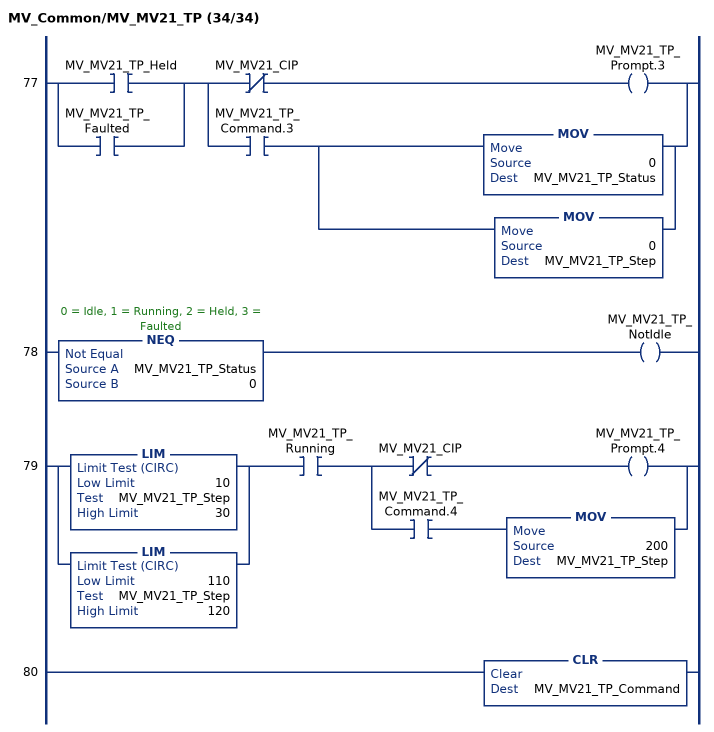
   77: [XIC(MV_MV21_TP_Held) ,XIC(MV_MV21_TP_Faulted) ][XIO(MV_MV21_CIP) OTE(MV_MV21_TP_Prompt.3) ,XIC(MV_MV21_TP_Command.3) [MOV(0,MV_MV21_TP_Status) ,MOV(0,MV_MV21_TP_Step) ] ];
   78: NEQ(MV_MV21_TP_Status,0)OTE(MV_MV21_TP_NotIdle);
   79: [LIM(10,MV_MV21_TP_Step,30) ,LIM(110,MV_MV21_TP_Step,120) ]XIC(MV_MV21_TP_Running)[XIO(MV_MV21_CIP) OTE(MV_MV21_TP_Prompt.4) ,XIC(MV_MV21_TP_Command.4) MOV(200,MV_MV21_TP_Step) ];
   80: CLR(MV_MV21_TP_Command);
END_ROUTINE

ROUTINE MV_MV22_TP   (* ladder *)
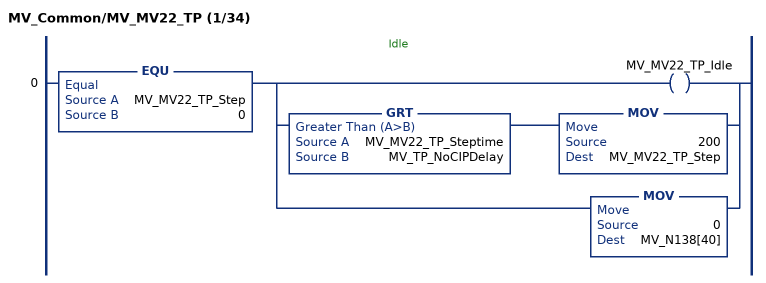
   // Idle
   0: EQU(MV_MV22_TP_Step,0)[OTE(MV_MV22_TP_Idle) ,GRT(MV_MV22_TP_Steptime,MV_TP_NoCIPDelay) MOV(200,MV_MV22_TP_Step) ,MOV(0,MV_N138[40]) ];
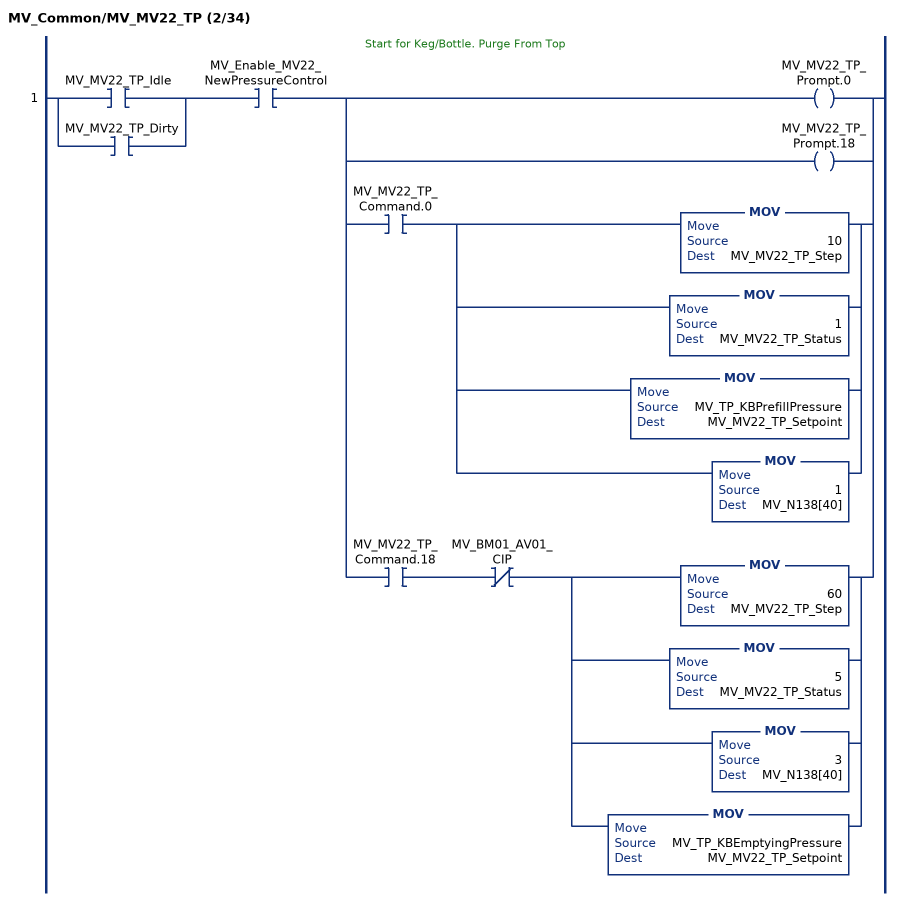
   // Start for Keg/Bottle. Purge From Top
   1: [XIC(MV_MV22_TP_Idle) ,XIC(MV_MV22_TP_Dirty) ]XIC(MV_Enable_MV22_NewPressureControl)[OTE(MV_MV22_TP_Prompt.0) ,OTE(MV_MV22_TP_Prompt.18) ,XIC(MV_MV22_TP_Command.0) [MOV(10,MV_MV22_TP_Step) ,MOV(1,MV_MV22_TP_Status) ,MOV(MV_TP_KBPrefillPressure,MV_MV22_TP_Setpoint) ,MOV(1,MV_N138[40]) ] ,XIC(MV_MV22_TP_Command.18) XIO(MV_BM01_AV01_CIP) [MOV(60,MV_MV22_TP_Step) ,MOV(5,MV_MV22_TP_Status) ,MOV(3,MV_N138[40]) ,MOV(MV_TP_KBEmptyingPressure,MV_MV22_TP_Setpoint) ] ];
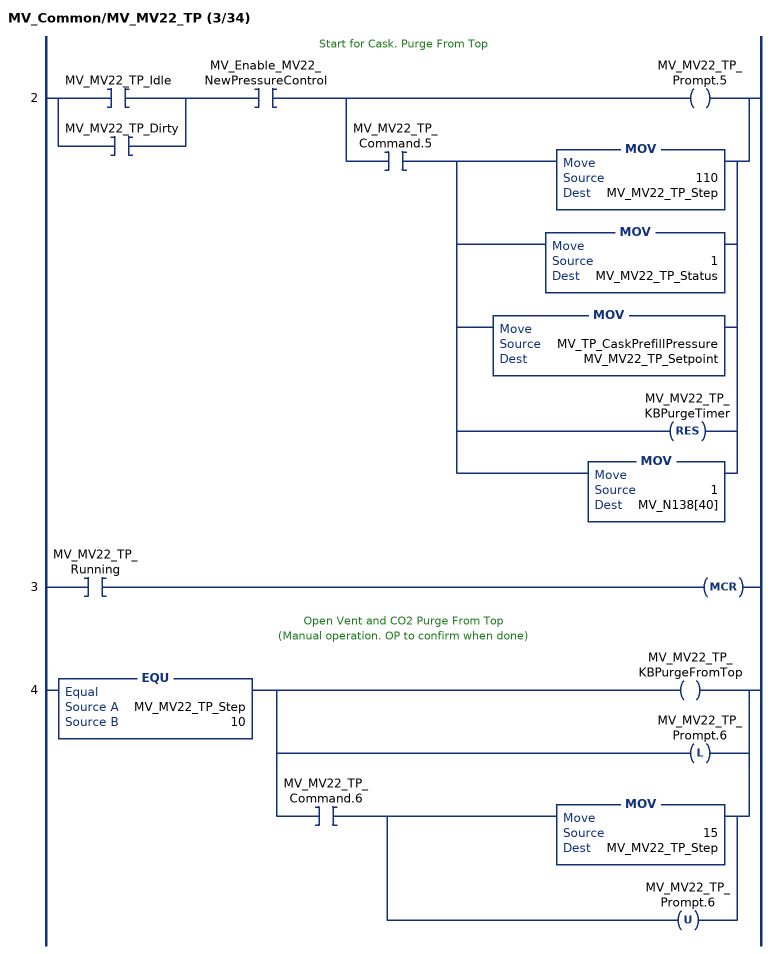
   // Start for Cask. Purge From Top
   2: [XIC(MV_MV22_TP_Idle) ,XIC(MV_MV22_TP_Dirty) ]XIC(MV_Enable_MV22_NewPressureControl)[OTE(MV_MV22_TP_Prompt.5) ,XIC(MV_MV22_TP_Command.5) [MOV(110,MV_MV22_TP_Step) ,MOV(1,MV_MV22_TP_Status) ,MOV(MV_TP_CaskPrefillPressure,MV_MV22_TP_Setpoint) ,RES(MV_MV22_TP_KBPurgeTimer) ,MOV(1,MV_N138[40]) ] ];
   3: XIC(MV_MV22_TP_Running)MCR();
   // Open Vent and CO2 Purge From Top
   // (Manual operation. OP to confirm when done)
   4: EQU(MV_MV22_TP_Step,10)[OTE(MV_MV22_TP_KBPurgeFromTop) ,OTL(MV_MV22_TP_Prompt.6) ,XIC(MV_MV22_TP_Command.6) [MOV(15,MV_MV22_TP_Step) ,OTU(MV_MV22_TP_Prompt.6) ] ];
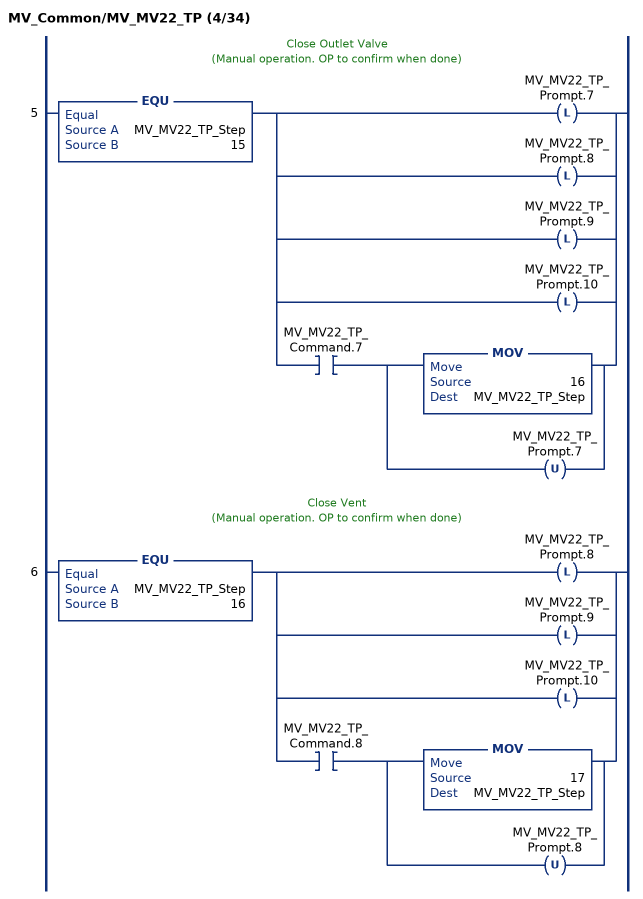
   // Close Outlet Valve
   // (Manual operation. OP to confirm when done)
   5: EQU(MV_MV22_TP_Step,15)[OTL(MV_MV22_TP_Prompt.7) ,OTL(MV_MV22_TP_Prompt.8) ,OTL(MV_MV22_TP_Prompt.9) ,OTL(MV_MV22_TP_Prompt.10) ,XIC(MV_MV22_TP_Command.7) [MOV(16,MV_MV22_TP_Step) ,OTU(MV_MV22_TP_Prompt.7) ] ];
   // Close Vent
   // (Manual operation. OP to confirm when done)
   6: EQU(MV_MV22_TP_Step,16)[OTL(MV_MV22_TP_Prompt.8) ,OTL(MV_MV22_TP_Prompt.9) ,OTL(MV_MV22_TP_Prompt.10) ,XIC(MV_MV22_TP_Command.8) [MOV(17,MV_MV22_TP_Step) ,OTU(MV_MV22_TP_Prompt.8) ] ];
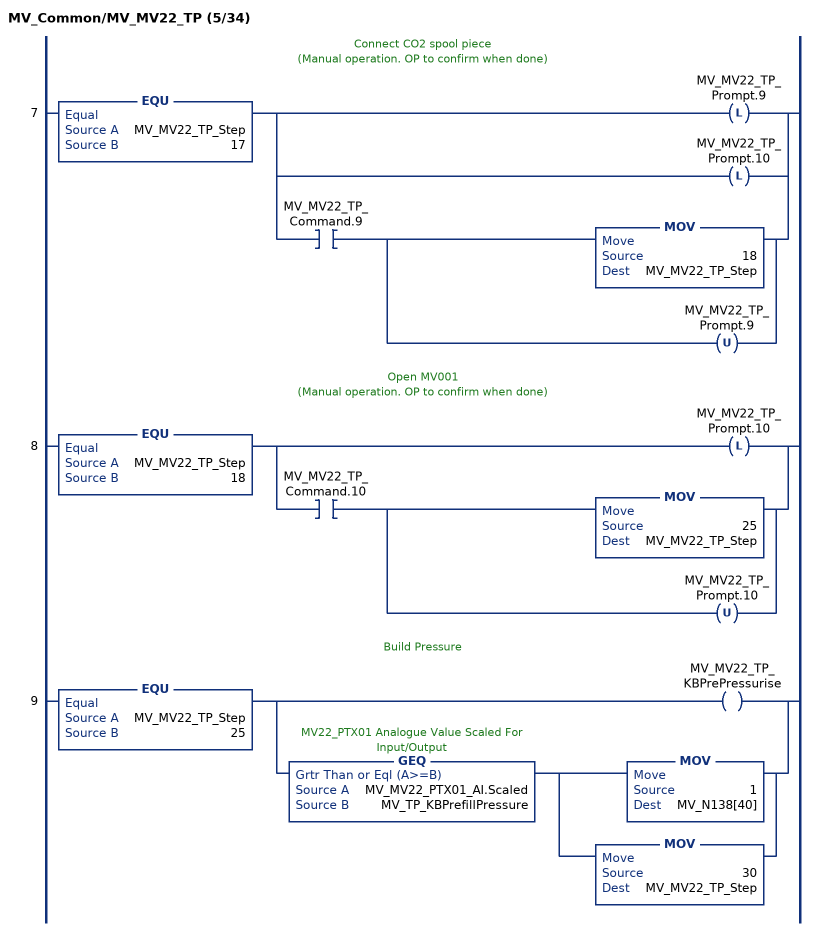
   // Connect CO2 spool piece
   // (Manual operation. OP to confirm when done)
   7: EQU(MV_MV22_TP_Step,17)[OTL(MV_MV22_TP_Prompt.9) ,OTL(MV_MV22_TP_Prompt.10) ,XIC(MV_MV22_TP_Command.9) [MOV(18,MV_MV22_TP_Step) ,OTU(MV_MV22_TP_Prompt.9) ] ];
   // Open MV001
   // (Manual operation. OP to confirm when done)
   8: EQU(MV_MV22_TP_Step,18)[OTL(MV_MV22_TP_Prompt.10) ,XIC(MV_MV22_TP_Command.10) [MOV(25,MV_MV22_TP_Step) ,OTU(MV_MV22_TP_Prompt.10) ] ];
   // Build Pressure
   9: EQU(MV_MV22_TP_Step,25)[OTE(MV_MV22_TP_KBPrePressurise) ,GEQ(MV_MV22_PTX01_AI.Scaled,MV_TP_KBPrefillPressure) [MOV(1,MV_N138[40]) ,MOV(30,MV_MV22_TP_Step) ] ];
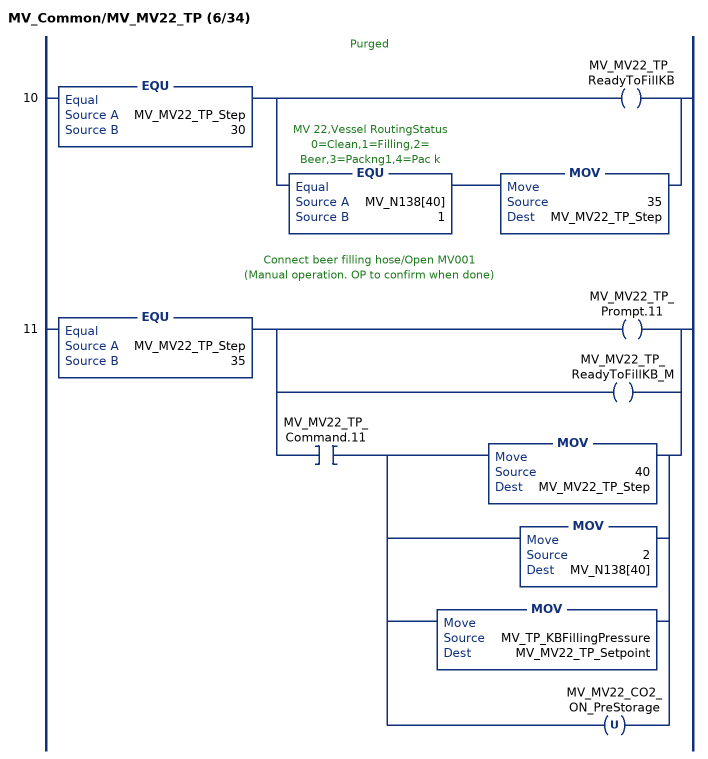
   // Purged
   10: EQU(MV_MV22_TP_Step,30)[OTE(MV_MV22_TP_ReadyToFillKB) ,EQU(MV_N138[40],1) MOV(35,MV_MV22_TP_Step) ];
   // Connect beer filling hose/Open MV001
   // (Manual operation. OP to confirm when done)
   11: EQU(MV_MV22_TP_Step,35)[OTE(MV_MV22_TP_Prompt.11) ,OTE(MV_MV22_TP_ReadyToFillKB_M) ,XIC(MV_MV22_TP_Command.11) [MOV(40,MV_MV22_TP_Step) ,MOV(2,MV_N138[40]) ,MOV(MV_TP_KBFillingPressure,MV_MV22_TP_Setpoint) ,OTU(MV_MV22_CO2_ON_PreStorage) ] ];
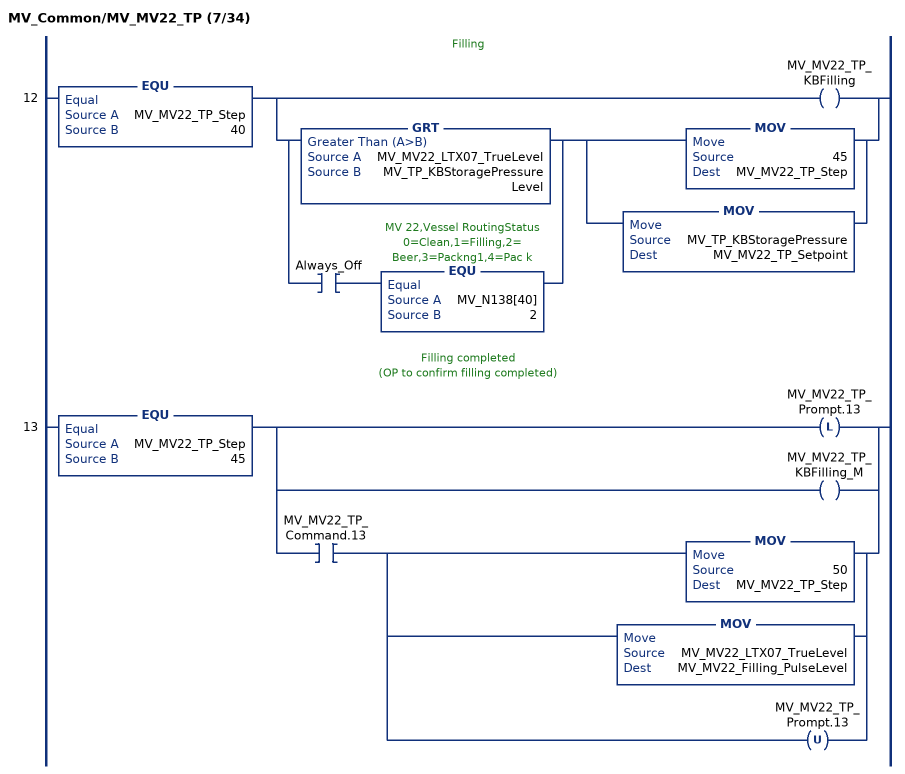
   // Filling
   12: EQU(MV_MV22_TP_Step,40)[OTE(MV_MV22_TP_KBFilling) ,[GRT(MV_MV22_LTX07_TrueLevel,MV_TP_KBStoragePressureLevel) ,XIC(Always_Off) EQU(MV_N138[40],2) ] [MOV(45,MV_MV22_TP_Step) ,MOV(MV_TP_KBStoragePressure,MV_MV22_TP_Setpoint) ] ];
   // Filling completed
   // (OP to confirm filling completed)
   13: EQU(MV_MV22_TP_Step,45)[OTL(MV_MV22_TP_Prompt.13) ,OTE(MV_MV22_TP_KBFilling_M) ,XIC(MV_MV22_TP_Command.13) [MOV(50,MV_MV22_TP_Step) ,MOV(MV_MV22_LTX07_TrueLevel,MV_MV22_Filling_PulseLevel) ,OTU(MV_MV22_TP_Prompt.13) ] ];
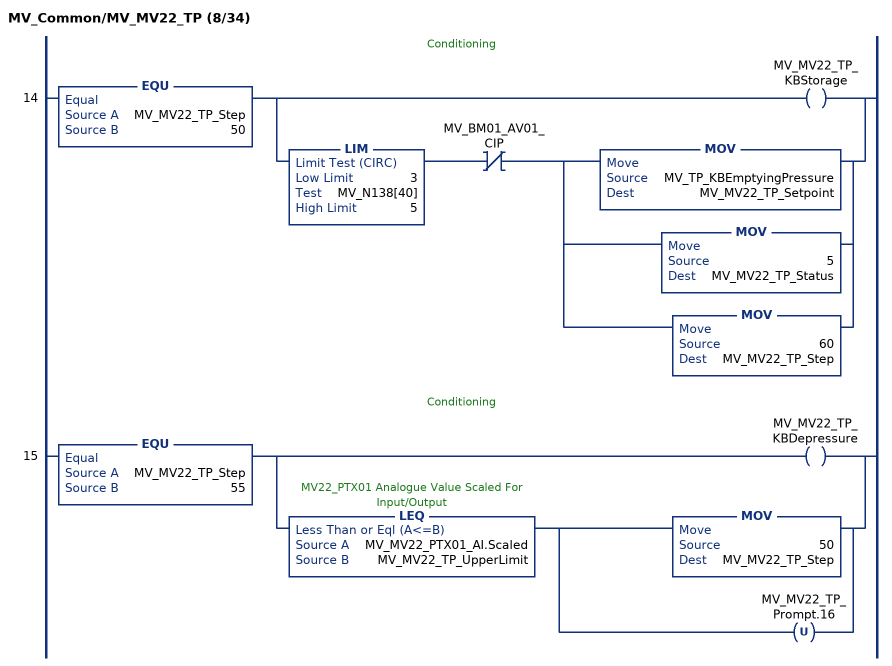
   // Conditioning
   14: EQU(MV_MV22_TP_Step,50)[OTE(MV_MV22_TP_KBStorage) ,LIM(3,MV_N138[40],5) XIO(MV_BM01_AV01_CIP) [MOV(MV_TP_KBEmptyingPressure,MV_MV22_TP_Setpoint) ,MOV(5,MV_MV22_TP_Status) ,MOV(60,MV_MV22_TP_Step) ] ];
   // Conditioning
   15: EQU(MV_MV22_TP_Step,55)[OTE(MV_MV22_TP_KBDepressure) ,LEQ(MV_MV22_PTX01_AI.Scaled,MV_MV22_TP_UpperLimit) [MOV(50,MV_MV22_TP_Step) ,OTU(MV_MV22_TP_Prompt.16) ] ];
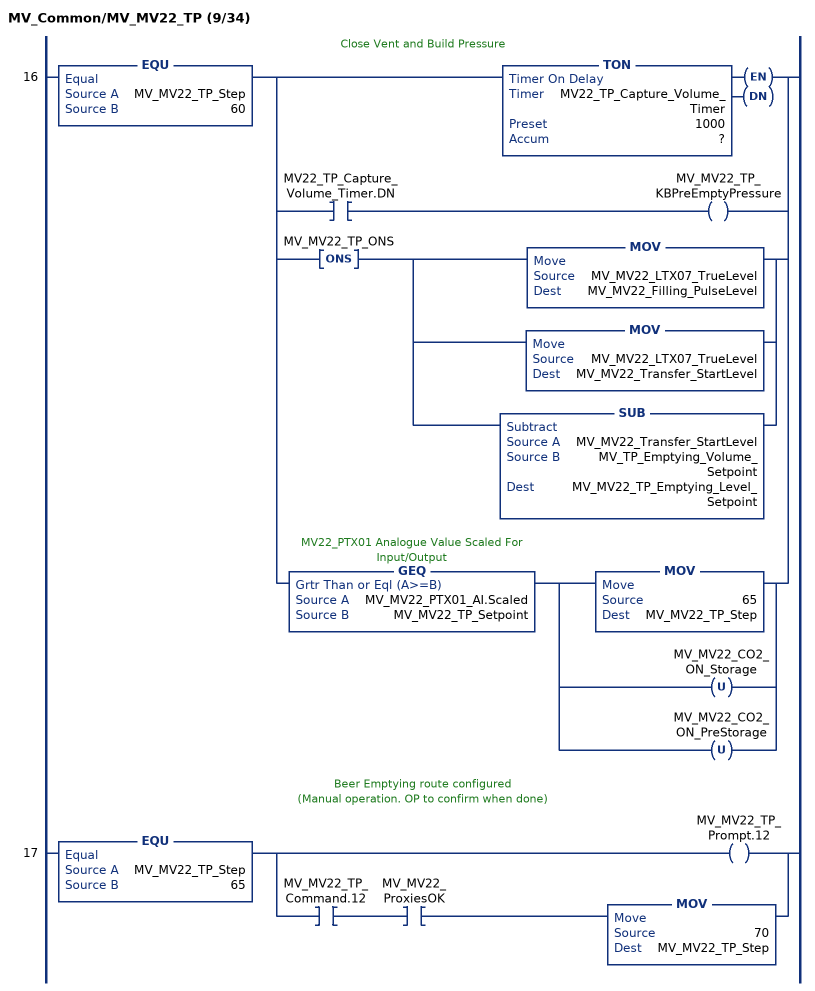
   // Close Vent and Build Pressure
   16: EQU(MV_MV22_TP_Step,60)[TON(MV22_TP_Capture_Volume_Timer,?,?) ,XIC(MV22_TP_Capture_Volume_Timer.DN) OTE(MV_MV22_TP_KBPreEmptyPressure) ,ONS(MV_MV22_TP_ONS) [MOV(MV_MV22_LTX07_TrueLevel,MV_MV22_Filling_PulseLevel) ,MOV(MV_MV22_LTX07_TrueLevel,MV_MV22_Transfer_StartLevel) ,SUB(MV_MV22_Transfer_StartLevel,MV_TP_Emptying_Volume_Setpoint,MV_MV22_TP_Emptying_Level_Setpoint) ] ,GEQ(MV_MV22_PTX01_AI.Scaled,MV_MV22_TP_Setpoint) [MOV(65,MV_MV22_TP_Step) ,OTU(MV_MV22_CO2_ON_Storage) ,OTU(MV_MV22_CO2_ON_PreStorage) ] ];
   // Beer Emptying route configured
   // (Manual operation. OP to confirm when done)
   17: EQU(MV_MV22_TP_Step,65)[OTE(MV_MV22_TP_Prompt.12) ,XIC(MV_MV22_TP_Command.12) XIC(MV_MV22_ProxiesOK) MOV(70,MV_MV22_TP_Step) ];
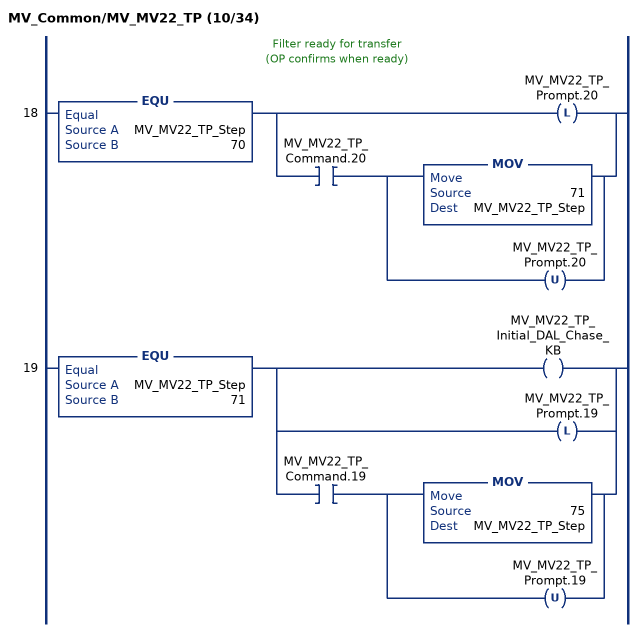
   // Filter ready for transfer
   // (OP confirms when ready)
   18: EQU(MV_MV22_TP_Step,70)[OTL(MV_MV22_TP_Prompt.20) ,XIC(MV_MV22_TP_Command.20) [MOV(71,MV_MV22_TP_Step) ,OTU(MV_MV22_TP_Prompt.20) ] ];
   19: EQU(MV_MV22_TP_Step,71)[OTE(MV_MV22_TP_Initial_DAL_Chase_KB) ,OTL(MV_MV22_TP_Prompt.19) ,XIC(MV_MV22_TP_Command.19) [MOV(75,MV_MV22_TP_Step) ,OTU(MV_MV22_TP_Prompt.19) ] ];
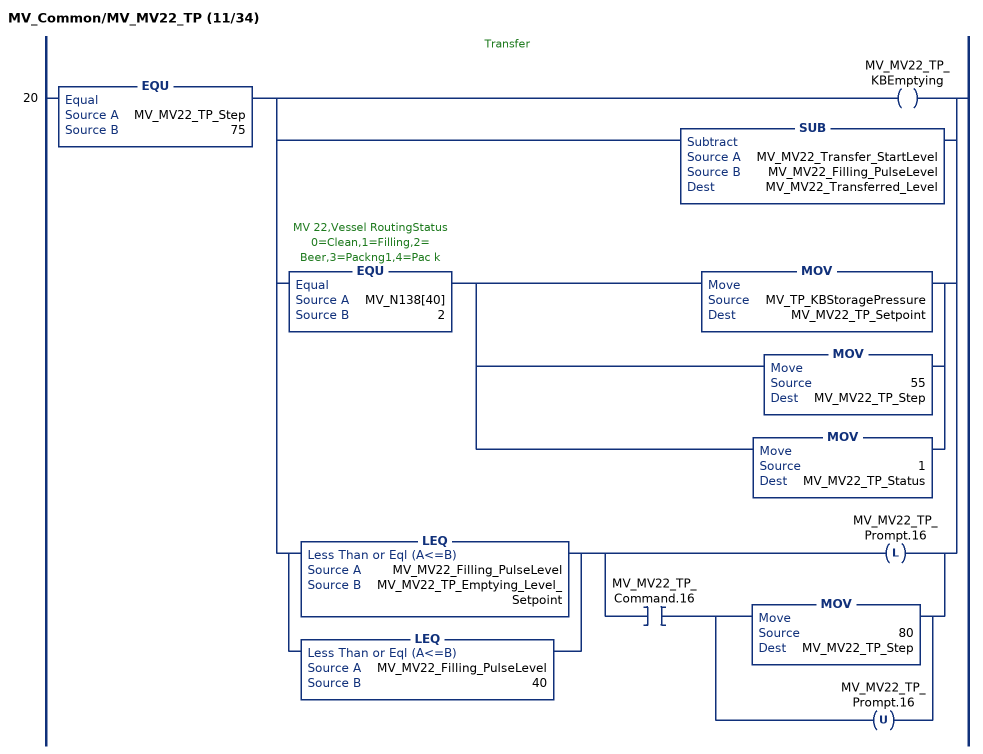
   // Transfer
   20: EQU(MV_MV22_TP_Step,75)[OTE(MV_MV22_TP_KBEmptying) ,SUB(MV_MV22_Transfer_StartLevel,MV_MV22_Filling_PulseLevel,MV_MV22_Transferred_Level) ,EQU(MV_N138[40],2) [MOV(MV_TP_KBStoragePressure,MV_MV22_TP_Setpoint) ,MOV(55,MV_MV22_TP_Step) ,MOV(1,MV_MV22_TP_Status) ] ,[LEQ(MV_MV22_Filling_PulseLevel,MV_MV22_TP_Emptying_Level_Setpoint) ,LEQ(MV_MV22_Filling_PulseLevel,40) ] [OTL(MV_MV22_TP_Prompt.16) ,XIC(MV_MV22_TP_Command.16) [MOV(80,MV_MV22_TP_Step) ,OTU(MV_MV22_TP_Prompt.16) ] ] ];
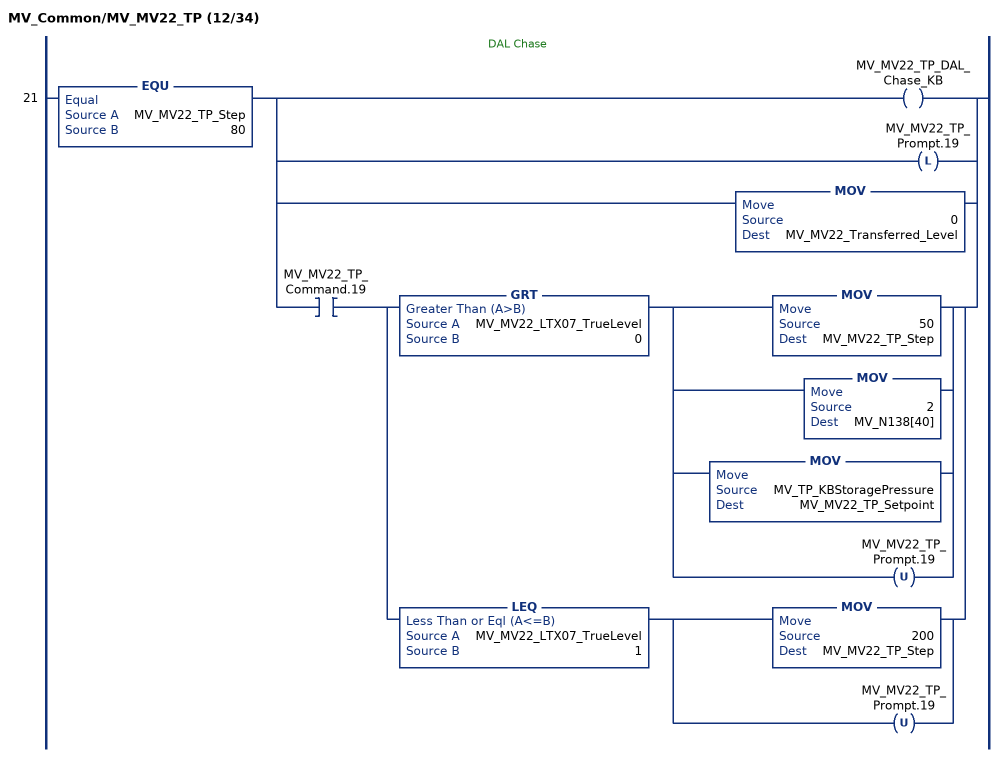
   // DAL Chase
   21: EQU(MV_MV22_TP_Step,80)[OTE(MV_MV22_TP_DAL_Chase_KB) ,OTL(MV_MV22_TP_Prompt.19) ,MOV(0,MV_MV22_Transferred_Level) ,XIC(MV_MV22_TP_Command.19) [GRT(MV_MV22_LTX07_TrueLevel,0) [MOV(50,MV_MV22_TP_Step) ,MOV(2,MV_N138[40]) ,MOV(MV_TP_KBStoragePressure,MV_MV22_TP_Setpoint) ,OTU(MV_MV22_TP_Prompt.19) ] ,LEQ(MV_MV22_LTX07_TrueLevel,1) [MOV(200,MV_MV22_TP_Step) ,OTU(MV_MV22_TP_Prompt.19) ] ] ];
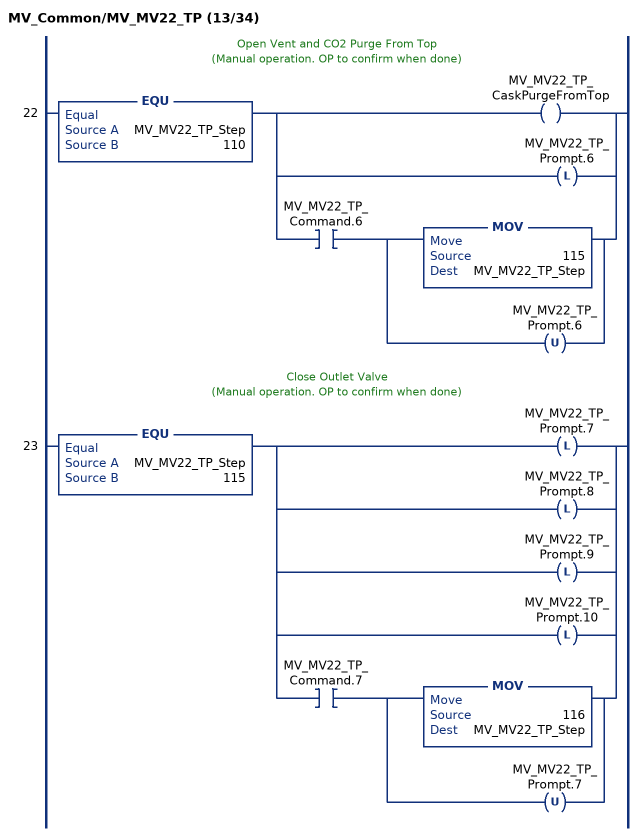
   // Open Vent and CO2 Purge From Top
   // (Manual operation. OP to confirm when done)
   22: EQU(MV_MV22_TP_Step,110)[OTE(MV_MV22_TP_CaskPurgeFromTop) ,OTL(MV_MV22_TP_Prompt.6) ,XIC(MV_MV22_TP_Command.6) [MOV(115,MV_MV22_TP_Step) ,OTU(MV_MV22_TP_Prompt.6) ] ];
   // Close Outlet Valve
   // (Manual operation. OP to confirm when done)
   23: EQU(MV_MV22_TP_Step,115)[OTL(MV_MV22_TP_Prompt.7) ,OTL(MV_MV22_TP_Prompt.8) ,OTL(MV_MV22_TP_Prompt.9) ,OTL(MV_MV22_TP_Prompt.10) ,XIC(MV_MV22_TP_Command.7) [MOV(116,MV_MV22_TP_Step) ,OTU(MV_MV22_TP_Prompt.7) ] ];
